(* Logix 5000 project; controller PLC_MCC1300_75F1 vendor 1 type 14 code 166 rev 32.11; software revision 32.04; part 57 of 83 *)
(* tags used below, declared in another part *)
   CM_AreaStackerToLine_JS1_Sync : CM_AreaStackerToLine;
   CM_ConveyorStackerToLine_JS1_Sync : CM_ConveyorStackerToLine;
   CM_DATA_Z410_Tx : UDT_PlateData_Convoy;
   CM_DATA_Z410_Tx_PH : DINT;
   CM_LineToAreaStacker_JS1 : CM_LineToAreaStacker;
   CM_LineToConveyorStacker_JS1 : CM_LineToConveyorStacker;
   CONST_dDest_Cullet : DINT;
   CONST_dDest_Stk : DINT;
   CONST_rgdDestMask : DINT[32];   // Destination Mask
   Convoy_SL_DATA_NULL : UDT_Convoy_SL;
   GP_CheckIdPlatePresent : GP_CheckIdPlatePresent;
   GP_CompactConvoy : GP_CompactConvoy;
   GP_ConvertDataToStacker : GP_ConvertDataToStacker;
   GP_OB_InitializeMain : GP_OB_Initialize;
   GP_RampSpace : GP_RampSpace;
   Gp_SpaceConvUtilities_V1 : GP_SpaceConvUtilities_V1;
   M311 : MAC_Conveyor;
   M311_Data : UDT_Convoy_SL;
   M311_SpaceConv_Utilities : SpaceConv_Utilities;
   M311M312_OffsetBaricentre_cmm : DINT;
   M312 : MAC_Conveyor_Single;
   M312_Data : UDT_Convoy_SL;
   M312_dSlowingSquaringQuote : DINT;
   M312_HMW : MAC_Conveyor_HMW;
   M312_M1_DR_IN_MAM : MOTION_INSTRUCTION;
   M312_SpaceConv_Utilities : SpaceConv_Utilities;
   M312_TON_Load : TIMER;
   M312_xEnableTractionRecovering : BOOL;
   M312_xLateralTractionRecovered : BOOL;
   M312_xPlateCullet : BOOL;
   M312_xSendCulletReqActive : BOOL;
   TMP_CenterLites : BOOL;
   TMP_d : DINT;
   TMP_dConveyorNumberForZoneCleaning : DINT;
   TMP_dDecelerationPositionEndConveyor : DINT;
   TMP_DistanceLateralSquaringToCenter : DINT;
   TMP_dOffsetLoadUnload_cmm : DINT;
   TMP_LiteAHeadY : DINT;
   TMP_LiteATailY : DINT;
   TMP_LiteBHeadY : DINT;
   TMP_LiteBTailY : DINT;
   TMP_rgxId : DINT[10];
   TMP_SquaringPosition : DINT;
   TMP_xConveyorInvolvedInCleaning : BOOL;
   TMP_xConveyorOfStartCleaning : BOOL;
   TMP_xCulletPresent : BOOL;
   TMP_xEnableLoadUnload : BOOL;
   TMP_xEnableZoneCleaning : BOOL;
   TMP_xLiteThisDestPresent : BOOL;
   x311PortraitMode : BOOL;
   xAlwaysOFF : BOOL;
   xAlwaysON : BOOL;
   xDebugOFF : BOOL;
   Z401 : MAC_Zone;
   Z401_HMR : MAC_Zone_HMR;
   Z401_HMW : MAC_Zone_HMW;
   Z401S_INPUT_xSafetyAreaPopup : BOOL;
(* MainProgram, continued *)

ROUTINE M312_Logic   (* ladder *)
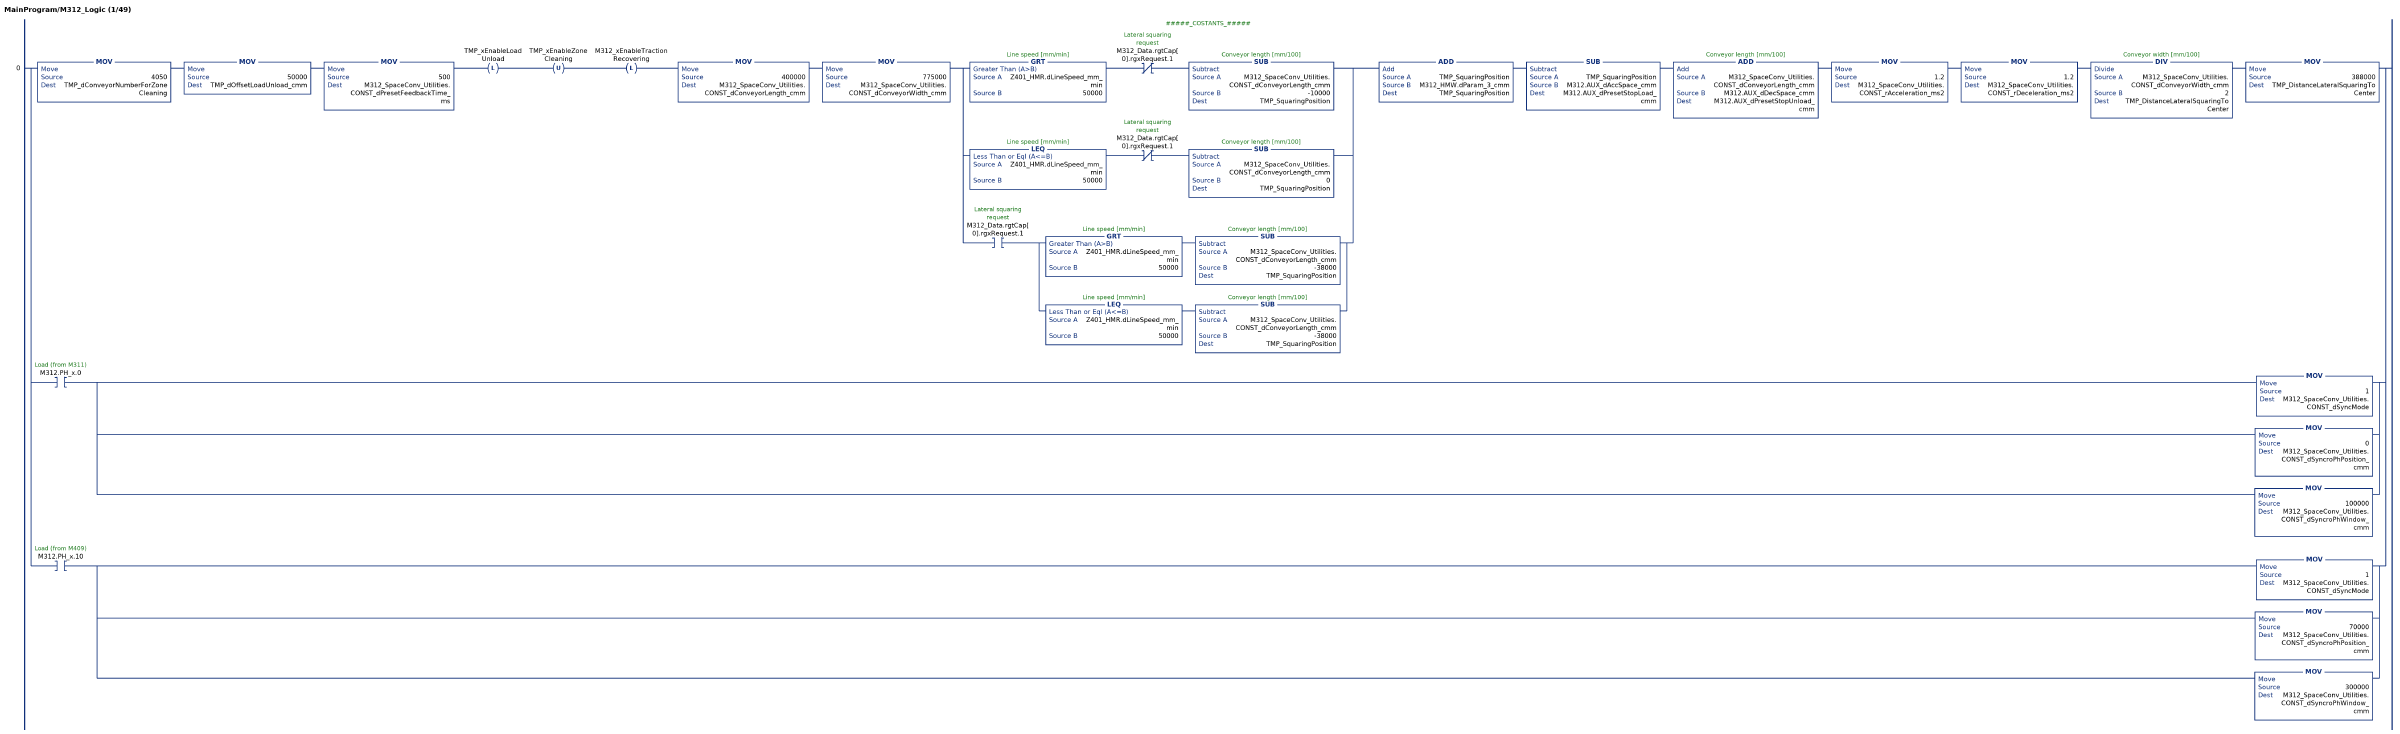
   // #####_COSTANTS_#####
   0: [MOV(4050,TMP_dConveyorNumberForZoneCleaning) MOV(50000,TMP_dOffsetLoadUnload_cmm) MOV(500,M312_SpaceConv_Utilities.CONST_dPresetFeedbackTime_ms) OTL(TMP_xEnableLoadUnload) OTU(TMP_xEnableZoneCleaning) OTL(M312_xEnableTractionRecovering) MOV(400000,M312_SpaceConv_Utilities.CONST_dConveyorLength_cmm) MOV(775000,M312_SpaceConv_Utilities.CONST_dConveyorWidth_cmm) [GRT(Z401_HMR.dLineSpeed_mm_min,50000) XIO(M312_Data.rgtCap[0].rgxRequest.1) SUB(M312_SpaceConv_Utilities.CONST_dConveyorLength_cmm,-10000,TMP_SquaringPosition) ,LEQ(Z401_HMR.dLineSpeed_mm_min,50000) XIO(M312_Data.rgtCap[0].rgxRequest.1) SUB(M312_SpaceConv_Utilities.CONST_dConveyorLength_cmm,0,TMP_SquaringPosition) ,XIC(M312_Data.rgtCap[0].rgxRequest.1) [GRT(Z401_HMR.dLineSpeed_mm_min,50000) SUB(M312_SpaceConv_Utilities.CONST_dConveyorLength_cmm,-38000,TMP_SquaringPosition) ,LEQ(Z401_HMR.dLineSpeed_mm_min,50000) SUB(M312_SpaceConv_Utilities.CONST_dConveyorLength_cmm,-38000,TMP_SquaringPosition) ] ] ADD(TMP_SquaringPosition,M312_HMW.dParam_3_cmm,TMP_SquaringPosition) SUB(TMP_SquaringPosition,M312.AUX_dAccSpace_cmm,M312.AUX_dPresetStopLoad_cmm) ADD(M312_SpaceConv_Utilities.CONST_dConveyorLength_cmm,M312.AUX_dDecSpace_cmm,M312.AUX_dPresetStopUnload_cmm) MOV(1.2,M312_SpaceConv_Utilities.CONST_rAcceleration_ms2) MOV(1.2,M312_SpaceConv_Utilities.CONST_rDeceleration_ms2) DIV(M312_SpaceConv_Utilities.CONST_dConveyorWidth_cmm,2,TMP_DistanceLateralSquaringToCenter) MOV(388000,TMP_DistanceLateralSquaringToCenter) ,[XIC(M312.PH_x.0) [MOV(1,M312_SpaceConv_Utilities.CONST_dSyncMode) ,MOV(0,M312_SpaceConv_Utilities.CONST_dSyncroPhPosition_cmm) ,MOV(100000,M312_SpaceConv_Utilities.CONST_dSyncroPhWindow_cmm) ] ,XIC(M312.PH_x.10) [MOV(1,M312_SpaceConv_Utilities.CONST_dSyncMode) ,MOV(70000,M312_SpaceConv_Utilities.CONST_dSyncroPhPosition_cmm) ,MOV(300000,M312_SpaceConv_Utilities.CONST_dSyncroPhWindow_cmm) ] ] ];
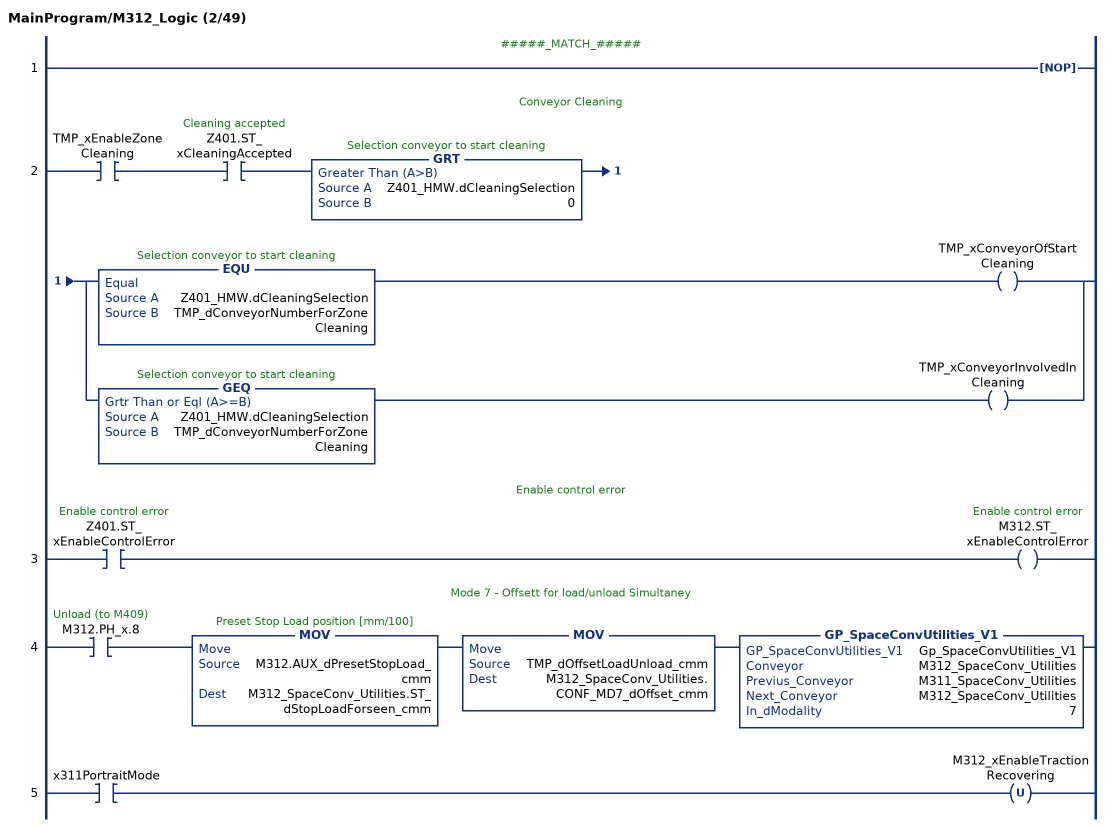
   // #####_MATCH_#####
   1: NOP();
   // Conveyor Cleaning
   2: XIC(TMP_xEnableZoneCleaning)XIC(Z401.ST_xCleaningAccepted)GRT(Z401_HMW.dCleaningSelection,0)[EQU(Z401_HMW.dCleaningSelection,TMP_dConveyorNumberForZoneCleaning) OTE(TMP_xConveyorOfStartCleaning) ,GEQ(Z401_HMW.dCleaningSelection,TMP_dConveyorNumberForZoneCleaning) OTE(TMP_xConveyorInvolvedInCleaning) ];
   // Enable control error
   3: XIC(Z401.ST_xEnableControlError)OTE(M312.ST_xEnableControlError);
   // Mode 7 - Offsett for load/unload Simultaney
   4: XIC(M312.PH_x.8)MOV(M312.AUX_dPresetStopLoad_cmm,M312_SpaceConv_Utilities.ST_dStopLoadForseen_cmm)MOV(TMP_dOffsetLoadUnload_cmm,M312_SpaceConv_Utilities.CONF_MD7_dOffset_cmm)GP_SpaceConvUtilities_V1(Gp_SpaceConvUtilities_V1,M312_SpaceConv_Utilities,M311_SpaceConv_Utilities,M312_SpaceConv_Utilities,7);
   5: XIC(x311PortraitMode)OTU(M312_xEnableTractionRecovering);
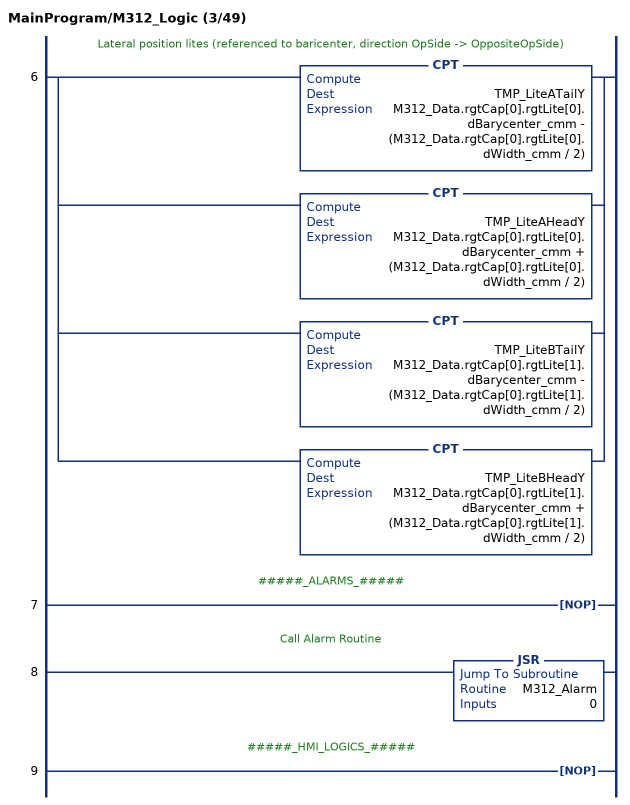
   // Lateral position lites (referenced to baricenter, direction OpSide -> OppositeOpSide)
   6: [CPT(TMP_LiteATailY,M312_Data.rgtCap[0].rgtLite[0].dBarycenter_cmm - (M312_Data.rgtCap[0].rgtLite[0].dWidth_cmm / 2)) ,CPT(TMP_LiteAHeadY,M312_Data.rgtCap[0].rgtLite[0].dBarycenter_cmm + (M312_Data.rgtCap[0].rgtLite[0].dWidth_cmm / 2)) ,CPT(TMP_LiteBTailY,M312_Data.rgtCap[0].rgtLite[1].dBarycenter_cmm - (M312_Data.rgtCap[0].rgtLite[1].dWidth_cmm / 2)) ,CPT(TMP_LiteBHeadY,M312_Data.rgtCap[0].rgtLite[1].dBarycenter_cmm + (M312_Data.rgtCap[0].rgtLite[1].dWidth_cmm / 2)) ];
   // #####_ALARMS_#####
   7: NOP();
   // Call Alarm Routine
   8: JSR(M312_Alarm,0);
   // #####_HMI_LOGICS_#####
   9: NOP();
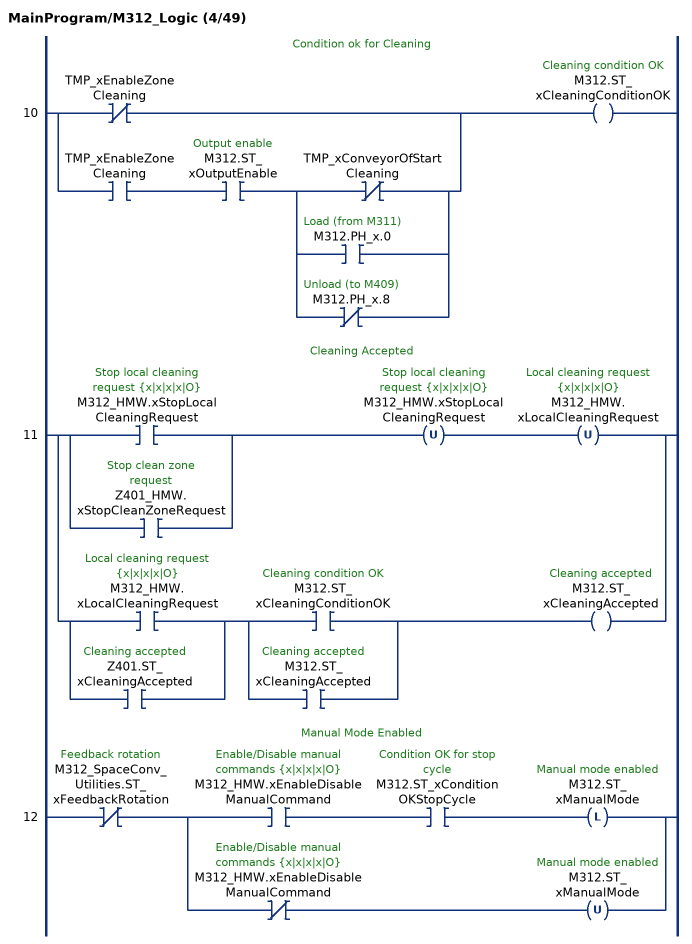
   // Condition ok for Cleaning
   10: [XIO(TMP_xEnableZoneCleaning) ,XIC(TMP_xEnableZoneCleaning) XIC(M312.ST_xOutputEnable) [XIO(TMP_xConveyorOfStartCleaning) ,XIC(M312.PH_x.0) ,XIO(M312.PH_x.8) ] ]OTE(M312.ST_xCleaningConditionOK);
   // Cleaning Accepted
   11: [[XIC(M312_HMW.xStopLocalCleaningRequest) ,XIC(Z401_HMW.xStopCleanZoneRequest) ] OTU(M312_HMW.xStopLocalCleaningRequest) OTU(M312_HMW.xLocalCleaningRequest) ,[XIC(M312_HMW.xLocalCleaningRequest) ,XIC(Z401.ST_xCleaningAccepted) ] [XIC(M312.ST_xCleaningConditionOK) ,XIC(M312.ST_xCleaningAccepted) ] OTE(M312.ST_xCleaningAccepted) ];
   // Manual Mode Enabled
   12: XIO(M312_SpaceConv_Utilities.ST_xFeedbackRotation)[XIC(M312_HMW.xEnableDisableManualCommand) XIC(M312.ST_xConditionOKStopCycle) OTL(M312.ST_xManualMode) ,XIO(M312_HMW.xEnableDisableManualCommand) OTU(M312.ST_xManualMode) ];
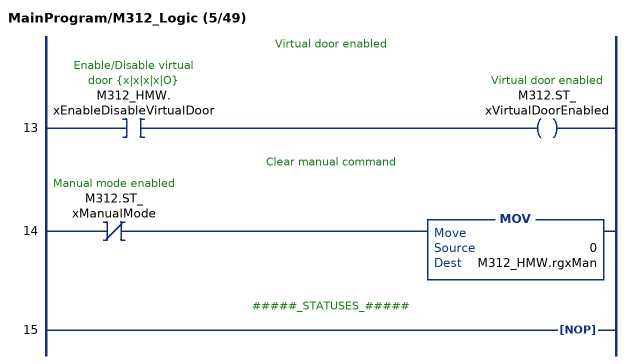
   // Virtual door enabled
   13: XIC(M312_HMW.xEnableDisableVirtualDoor)OTE(M312.ST_xVirtualDoorEnabled);
   // Clear manual command
   14: XIO(M312.ST_xManualMode)MOV(0,M312_HMW.rgxMan);
   // #####_STATUSES_#####
   15: NOP();
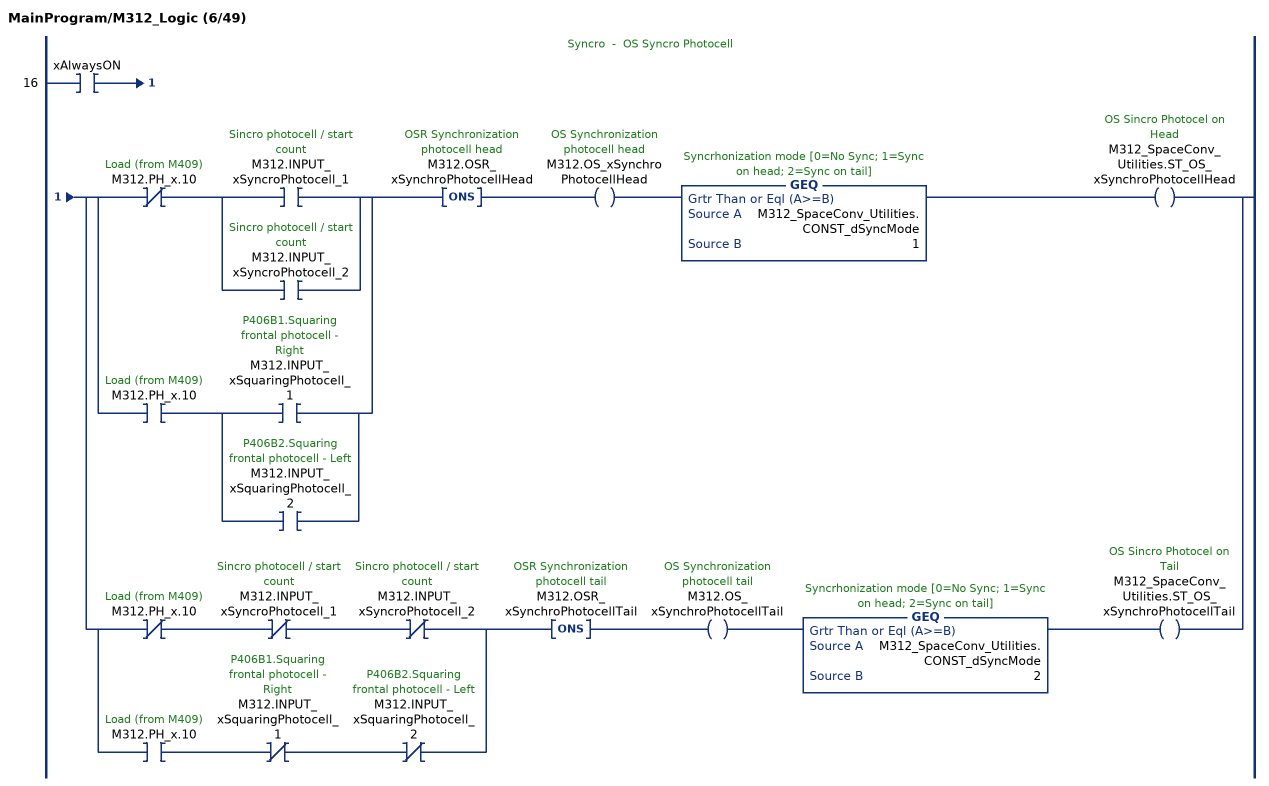
   // Syncro  -  OS Syncro Photocell
   16: XIC(xAlwaysON)[[XIO(M312.PH_x.10) [XIC(M312.INPUT_xSyncroPhotocell_1) ,XIC(M312.INPUT_xSyncroPhotocell_2) ] ,XIC(M312.PH_x.10) [XIC(M312.INPUT_xSquaringPhotocell_1) ,XIC(M312.INPUT_xSquaringPhotocell_2) ] ] ONS(M312.OSR_xSynchroPhotocellHead) OTE(M312.OS_xSynchroPhotocellHead) GEQ(M312_SpaceConv_Utilities.CONST_dSyncMode,1) OTE(M312_SpaceConv_Utilities.ST_OS_xSynchroPhotocellHead) ,[XIO(M312.PH_x.10) XIO(M312.INPUT_xSyncroPhotocell_1) XIO(M312.INPUT_xSyncroPhotocell_2) ,XIC(M312.PH_x.10) XIO(M312.INPUT_xSquaringPhotocell_1) XIO(M312.INPUT_xSquaringPhotocell_2) ] ONS(M312.OSR_xSynchroPhotocellTail) OTE(M312.OS_xSynchroPhotocellTail) GEQ(M312_SpaceConv_Utilities.CONST_dSyncMode,2) OTE(M312_SpaceConv_Utilities.ST_OS_xSynchroPhotocellTail) ];
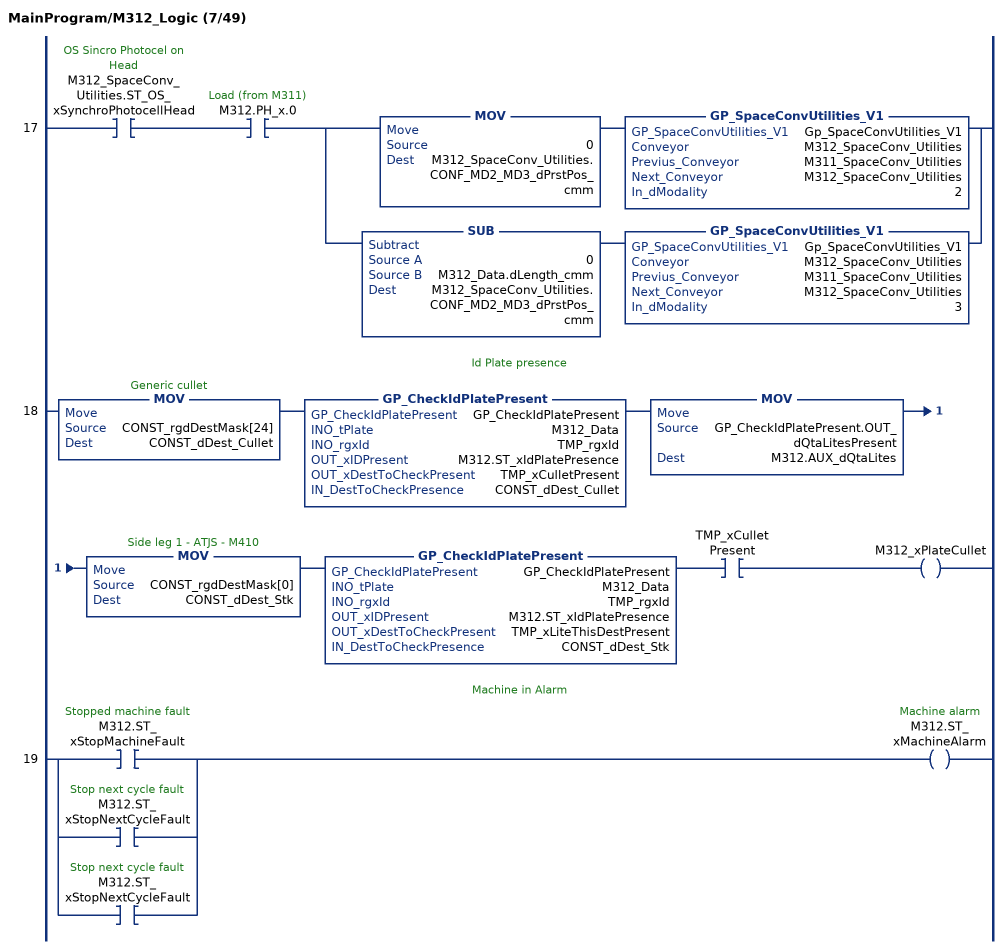
   17: XIC(M312_SpaceConv_Utilities.ST_OS_xSynchroPhotocellHead)XIC(M312.PH_x.0)[MOV(0,M312_SpaceConv_Utilities.CONF_MD2_MD3_dPrstPos_cmm) GP_SpaceConvUtilities_V1(Gp_SpaceConvUtilities_V1,M312_SpaceConv_Utilities,M311_SpaceConv_Utilities,M312_SpaceConv_Utilities,2) ,SUB(0,M312_Data.dLength_cmm,M312_SpaceConv_Utilities.CONF_MD2_MD3_dPrstPos_cmm) GP_SpaceConvUtilities_V1(Gp_SpaceConvUtilities_V1,M312_SpaceConv_Utilities,M311_SpaceConv_Utilities,M312_SpaceConv_Utilities,3) ];
   // Id Plate presence
   18: MOV(CONST_rgdDestMask[24],CONST_dDest_Cullet)GP_CheckIdPlatePresent(GP_CheckIdPlatePresent,M312_Data,TMP_rgxId,M312.ST_xIdPlatePresence,TMP_xCulletPresent,CONST_dDest_Cullet)MOV(GP_CheckIdPlatePresent.OUT_dQtaLitesPresent,M312.AUX_dQtaLites)MOV(CONST_rgdDestMask[0],CONST_dDest_Stk)GP_CheckIdPlatePresent(GP_CheckIdPlatePresent,M312_Data,TMP_rgxId,M312.ST_xIdPlatePresence,TMP_xLiteThisDestPresent,CONST_dDest_Stk)XIC(TMP_xCulletPresent)OTE(M312_xPlateCullet);
   // Machine in Alarm
   19: [XIC(M312.ST_xStopMachineFault) ,XIC(M312.ST_xStopNextCycleFault) ,XIC(M312.ST_xStopNextCycleFault) ]OTE(M312.ST_xMachineAlarm);
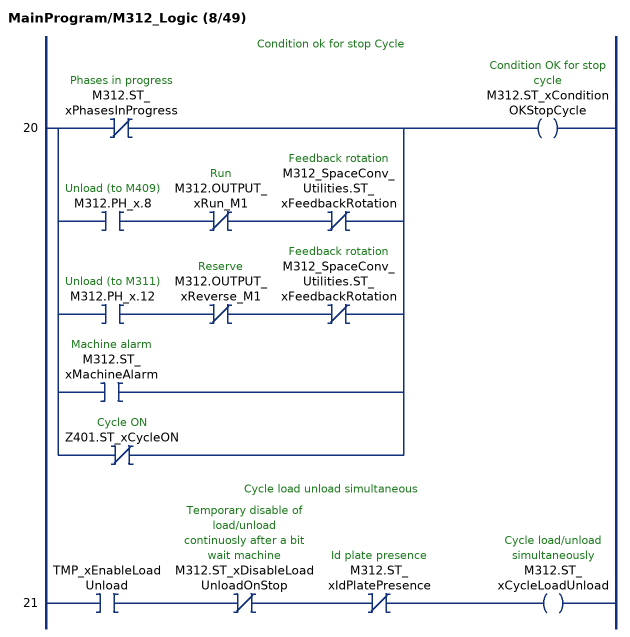
   // Condition ok for stop Cycle
   20: [XIO(M312.ST_xPhasesInProgress) ,XIC(M312.PH_x.8) XIO(M312.OUTPUT_xRun_M1) XIO(M312_SpaceConv_Utilities.ST_xFeedbackRotation) ,XIC(M312.PH_x.12) XIO(M312.OUTPUT_xReverse_M1) XIO(M312_SpaceConv_Utilities.ST_xFeedbackRotation) ,XIC(M312.ST_xMachineAlarm) ,XIO(Z401.ST_xCycleON) ]OTE(M312.ST_xConditionOKStopCycle);
   // Cycle load unload simultaneous
   21: XIC(TMP_xEnableLoadUnload)XIO(M312.ST_xDisableLoadUnloadOnStop)XIO(M312.ST_xIdPlatePresence)OTE(M312.ST_xCycleLoadUnload);
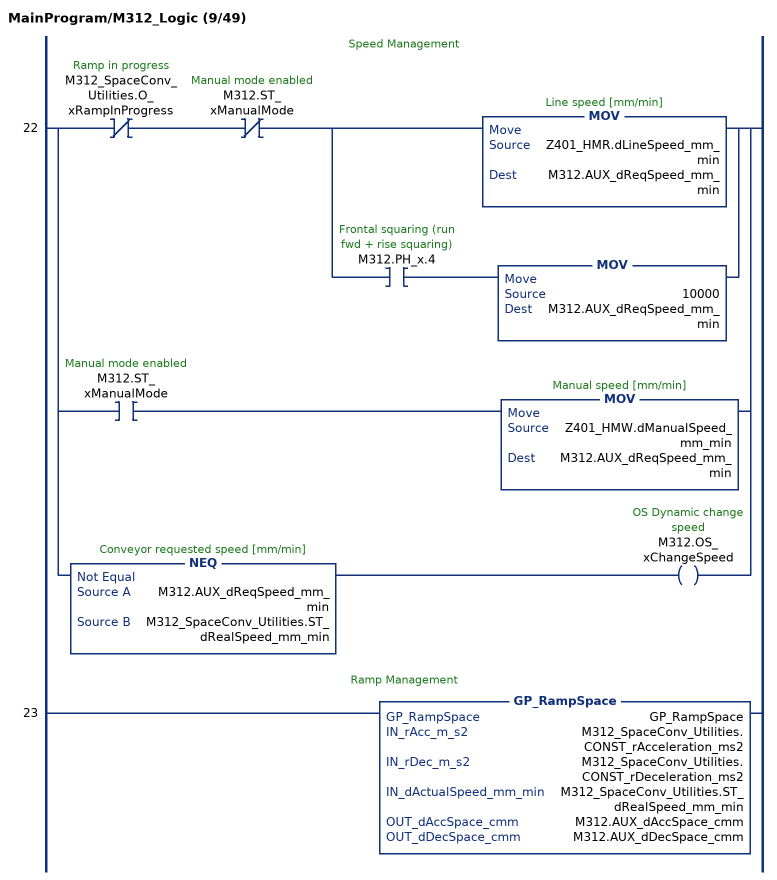
   // Speed Management
   22: [XIO(M312_SpaceConv_Utilities.O_xRampInProgress) XIO(M312.ST_xManualMode) [MOV(Z401_HMR.dLineSpeed_mm_min,M312.AUX_dReqSpeed_mm_min) ,XIC(M312.PH_x.4) MOV(10000,M312.AUX_dReqSpeed_mm_min) ] ,XIC(M312.ST_xManualMode) MOV(Z401_HMW.dManualSpeed_mm_min,M312.AUX_dReqSpeed_mm_min) ,NEQ(M312.AUX_dReqSpeed_mm_min,M312_SpaceConv_Utilities.ST_dRealSpeed_mm_min) OTE(M312.OS_xChangeSpeed) ];
   // Ramp Management
   23: GP_RampSpace(GP_RampSpace,M312_SpaceConv_Utilities.CONST_rAcceleration_ms2,M312_SpaceConv_Utilities.CONST_rDeceleration_ms2,M312_SpaceConv_Utilities.ST_dRealSpeed_mm_min,M312.AUX_dAccSpace_cmm,M312.AUX_dDecSpace_cmm);
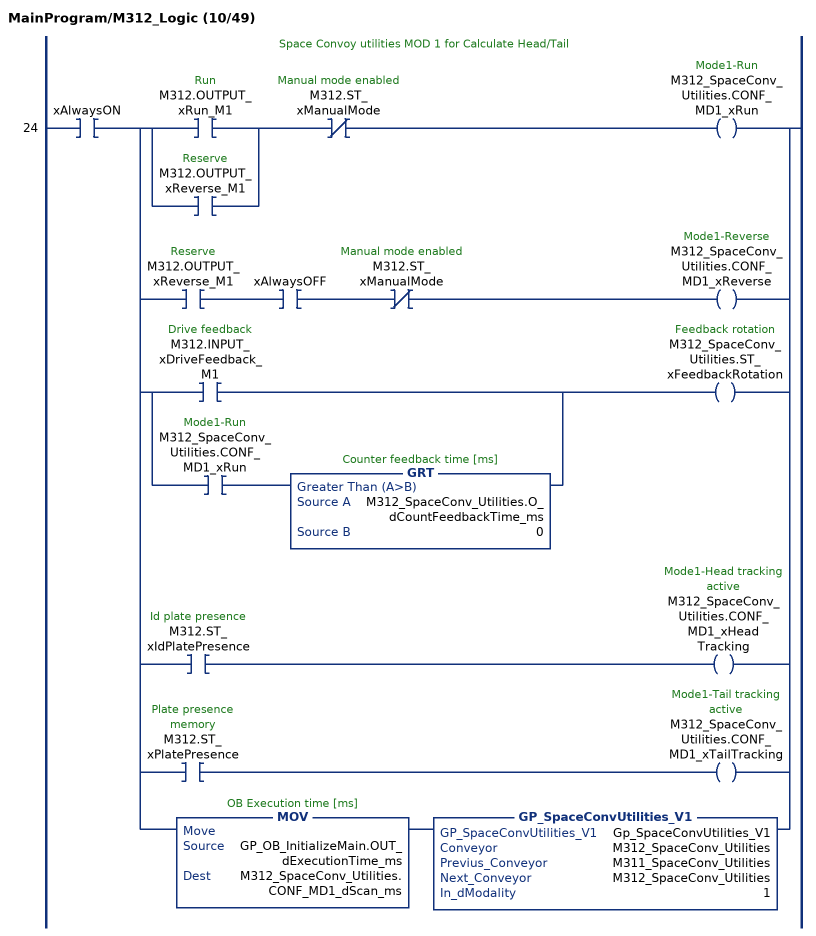
   // Space Convoy utilities MOD 1 for Calculate Head/Tail
   24: XIC(xAlwaysON)[[XIC(M312.OUTPUT_xRun_M1) ,XIC(M312.OUTPUT_xReverse_M1) ] XIO(M312.ST_xManualMode) OTE(M312_SpaceConv_Utilities.CONF_MD1_xRun) ,XIC(M312.OUTPUT_xReverse_M1) XIC(xAlwaysOFF) XIO(M312.ST_xManualMode) OTE(M312_SpaceConv_Utilities.CONF_MD1_xReverse) ,[XIC(M312.INPUT_xDriveFeedback_M1) ,XIC(M312_SpaceConv_Utilities.CONF_MD1_xRun) GRT(M312_SpaceConv_Utilities.O_dCountFeedbackTime_ms,0) ] OTE(M312_SpaceConv_Utilities.ST_xFeedbackRotation) ,XIC(M312.ST_xIdPlatePresence) OTE(M312_SpaceConv_Utilities.CONF_MD1_xHeadTracking) ,XIC(M312.ST_xPlatePresence) OTE(M312_SpaceConv_Utilities.CONF_MD1_xTailTracking) ,MOV(GP_OB_InitializeMain.OUT_dExecutionTime_ms,M312_SpaceConv_Utilities.CONF_MD1_dScan_ms) GP_SpaceConvUtilities_V1(Gp_SpaceConvUtilities_V1,M312_SpaceConv_Utilities,M311_SpaceConv_Utilities,M312_SpaceConv_Utilities,1) ];
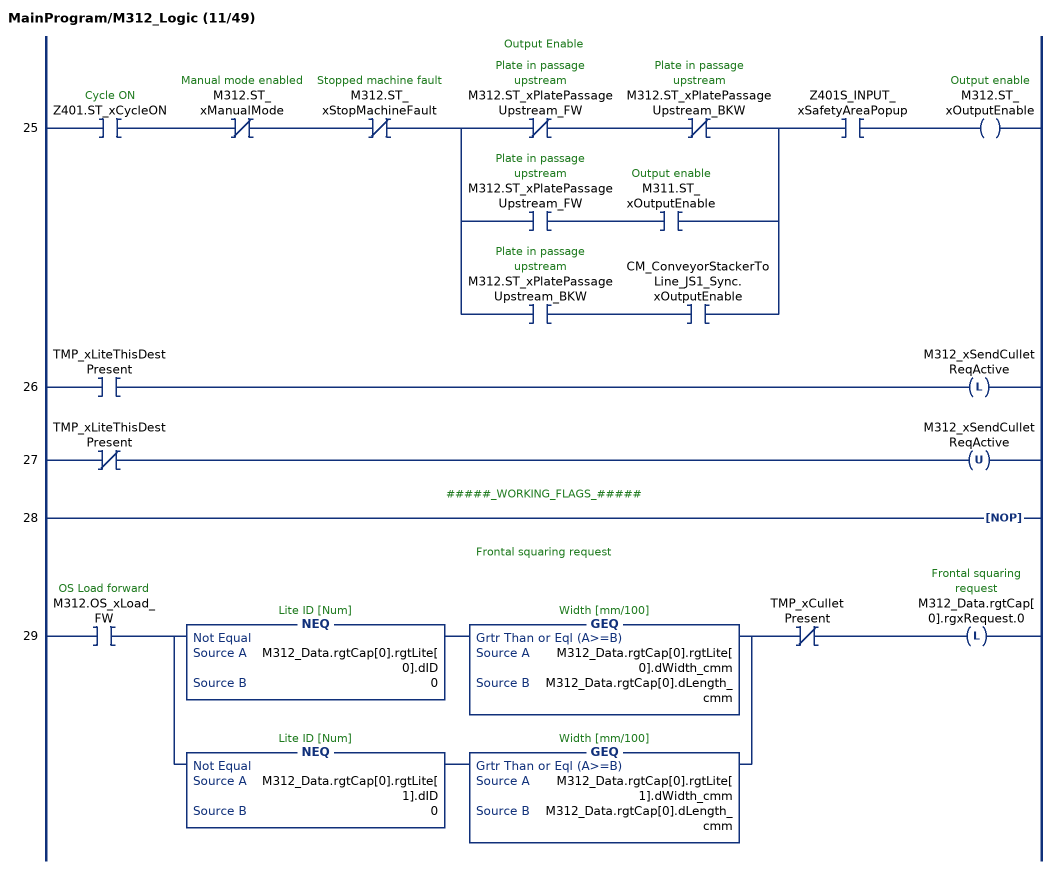
   // Output Enable
   25: XIC(Z401.ST_xCycleON)XIO(M312.ST_xManualMode)XIO(M312.ST_xStopMachineFault)[XIO(M312.ST_xPlatePassageUpstream_FW) XIO(M312.ST_xPlatePassageUpstream_BKW) ,XIC(M312.ST_xPlatePassageUpstream_FW) XIC(M311.ST_xOutputEnable) ,XIC(M312.ST_xPlatePassageUpstream_BKW) XIC(CM_ConveyorStackerToLine_JS1_Sync.xOutputEnable) ]XIC(Z401S_INPUT_xSafetyAreaPopup)OTE(M312.ST_xOutputEnable);
   26: XIC(TMP_xLiteThisDestPresent)OTL(M312_xSendCulletReqActive);
   27: XIO(TMP_xLiteThisDestPresent)OTU(M312_xSendCulletReqActive);
   // #####_WORKING_FLAGS_#####
   28: NOP();
   // Frontal squaring request
   29: XIC(M312.OS_xLoad_FW)[NEQ(M312_Data.rgtCap[0].rgtLite[0].dID,0) GEQ(M312_Data.rgtCap[0].rgtLite[0].dWidth_cmm,M312_Data.rgtCap[0].dLength_cmm) ,NEQ(M312_Data.rgtCap[0].rgtLite[1].dID,0) GEQ(M312_Data.rgtCap[0].rgtLite[1].dWidth_cmm,M312_Data.rgtCap[0].dLength_cmm) ]XIO(TMP_xCulletPresent)OTL(M312_Data.rgtCap[0].rgxRequest.0);